screen "05-Outputs1" 480x272, template "Main_Template"
   on GenerateScreen: SetTag("DB005-HMI_Data_iScreen_Number", 5)
   TextField "TextField_ScreenName" at 76,46 size 328x30; Text 'PLC DIGITAL OUTPUTS - 1of3'
   TextField "TextField_BankLetter" at 412,50 size 64x23; Text 'BANK A'
   Button "Button_Next" at 384,227 size 92x40; TextOff 'NEXT'
      on Press: ActivateScreen("06-Outputs2", 0)
   Group "Group_DQ0.0" at 18,83 size 97x62; TextList "ON/OFF"
   Group "Group_DQ0.1" at 132,83 size 97x62; TextList "ON/OFF"
   Group "Group_DQ0.2" at 247,83 size 97x62; TextList "ON/OFF"
   Group "Group_DQ0.3" at 362,83 size 97x62; TextList "ON/OFF"
   Group "Group_DQ0.4" at 18,154 size 97x62; TextList "ON/OFF"
   Group "Group_DQ0.5" at 132,154 size 97x62; TextList "ON/OFF"
   Group "Group_DQ0.6" at 247,154 size 97x62; TextList "ON/OFF"
   Group "Group_DQ0.7" at 362,154 size 97x62; TextList "ON/OFF"
   Rectangle "Rectangle_DQ0.0" at 18,83 size 97x62
      Appearance <- "DB001-PLC_I/O_Outputs_xDQ0.0"
   TextField "Text field_DQ0.0" at 44,83 size 46x19; Text 'DQ 0.0'
   Button "Button_DQ0.0" at 30,105 size 73x32; TextOff 'Text'; TextList "ON/OFF"
      on Press: InvertBit("DB001-PLC_I/O_Outputs_xDQ0.0")
      ProcessValue <- "DB001-PLC_I/O_Outputs_xDQ0.0"
   Rectangle "Rectangle_DQ0.1" at 132,83 size 97x62
      Appearance <- "DB001-PLC_I/O_Outputs_xDQ0.1"
   TextField "Text field_DQ0.1" at 158,83 size 46x19; Text 'DQ 0.1'
   Button "Button_DQ0.1" at 144,105 size 73x32; TextOff 'Text'; TextList "ON/OFF"
      on Press: InvertBit("DB001-PLC_I/O_Outputs_xDQ0.1")
      ProcessValue <- "DB001-PLC_I/O_Outputs_xDQ0.1"
   Rectangle "Rectangle_DQ0.2" at 247,83 size 97x62
      Appearance <- "DB001-PLC_I/O_Outputs_xDQ0.2"
   TextField "Text field_DQ0.2" at 273,83 size 46x19; Text 'DQ 0.2'
   Button "Button_DQ0.2" at 259,105 size 73x32; TextOff 'Text'; TextList "ON/OFF"
      on Press: InvertBit("DB001-PLC_I/O_Outputs_xDQ0.2")
      ProcessValue <- "DB001-PLC_I/O_Outputs_xDQ0.2"
   Rectangle "Rectangle_DQ0.3" at 362,83 size 97x62
      Appearance <- "DB001-PLC_I/O_Outputs_xDQ0.3"
   TextField "Text field_DQ0.3" at 388,83 size 46x19; Text 'DQ 0.3'
   Button "Button_DQ0.3" at 374,105 size 73x32; TextOff 'Text'; TextList "ON/OFF"
      on Press: InvertBit("DB001-PLC_I/O_Outputs_xDQ0.3")
      ProcessValue <- "DB001-PLC_I/O_Outputs_xDQ0.3"
   Rectangle "Rectangle_DQ0.4" at 18,154 size 97x62
      Appearance <- "DB001-PLC_I/O_Outputs_xDQ0.4"
   TextField "Text field_DQ0.4" at 44,154 size 46x19; Text 'DQ 0.4'
   Button "Button_DQ0.4" at 30,176 size 73x32; TextOff 'Text'; TextList "ON/OFF"
      on Press: InvertBit("DB001-PLC_I/O_Outputs_xDQ0.4")
      ProcessValue <- "DB001-PLC_I/O_Outputs_xDQ0.4"
   Rectangle "Rectangle_DQ0.5" at 132,154 size 97x62
      Appearance <- "DB001-PLC_I/O_Outputs_xDQ0.5"
   TextField "Text field_DQ0.5" at 158,154 size 46x19; Text 'DQ 0.5'
   Button "Button_DQ0.5" at 144,176 size 73x32; TextOff 'Text'; TextList "ON/OFF"
      on Press: InvertBit("DB001-PLC_I/O_Outputs_xDQ0.5")
      ProcessValue <- "DB001-PLC_I/O_Outputs_xDQ0.5"
   Rectangle "Rectangle_DQ0.6" at 247,154 size 97x62
      Appearance <- "DB001-PLC_I/O_Outputs_xDQ0.6"
   TextField "Text field_DQ0.6" at 273,154 size 46x19; Text 'DQ 0.6'
   Button "Button_DQ0.6" at 259,176 size 73x32; TextOff 'Text'; TextList "ON/OFF"
      on Press: InvertBit("DB001-PLC_I/O_Outputs_xDQ0.6")
      ProcessValue <- "DB001-PLC_I/O_Outputs_xDQ0.6"
   Rectangle "Rectangle_DQ0.7" at 362,154 size 97x62
      Appearance <- "DB001-PLC_I/O_Outputs_xDQ0.7"
   TextField "Text field_DQ0.7" at 388,154 size 46x19; Text 'DQ 0.7'
   Button "Button_DQ0.7" at 374,176 size 73x32; TextOff 'Text'; TextList "ON/OFF"
      on Press: InvertBit("DB001-PLC_I/O_Outputs_xDQ0.7")
      ProcessValue <- "DB001-PLC_I/O_Outputs_xDQ0.7"

screen "08-AnalogI/O" 480x272, template "Main_Template"
   on GenerateScreen: SetTag("DB005-HMI_Data_iScreen_Number", 8)
   Button "Button_Back" at 384,227 size 92x40; TextOff 'BACK'
      on Press: function_efd93a16()
   TextField "TextField_ScreenName" at 65,46 size 351x30; Text 'PLC ANALOG INPUTS/OUTPUTS'
   Group "Group_A0" at 244,76 size 229x145; FormatPattern 9999
   Group "Group_A1" at 8,76 size 229x145; FormatPattern 9999
   TextField "Text field_A0" at 291,77 size 127x21; Text 'Analog AI-0 & AQ-0'
   TextField "Text field_A0_Input" at 279,98 size 42x17; Text 'INPUT'
   TextField "Text field_A0_Instruction" at 256,115 size 86x34; Text 'Use the connected potentiometer to change the input voltage.'
   TextField "Text field_A0_Voltage" at 280,149 size 41x14; Text 'VOLTAGE:'
   IOField "I/O field_A0_Voltage" at 281,162 size 42x21; FormatPattern 99.99; Unit  V
      ProcessValue <- "DB001-PLC_I/O_Inputs_rAI0.0_Scaled"
   TextField "Text field_A0_InRAW" at 289,181 size 24x14; Text 'RAW:'
   IOField "I/O field_A0_RAW" at 283,193 size 37x21; FormatPattern 99999
      ProcessValue <- "AI0.0"
   TextField "Text field_A0_Output" at 389,98 size 52x17; Text 'OUTPUT'
   TextField "Text field_A0_mA" at 381,127 size 19x14; Text 'mA:'
   IOField "I/O field_A0_mA" at 365,140 size 51x21; FormatPattern 99.99; Unit  mA
      ProcessValue <- "DB001-PLC_I/O_Outputs_rAQ0.0_Scaled"
   TextField "Text field_A0_OutRAW" at 379,167 size 24x14; Text 'RAW:'
   IOField "I/O field_A0_OutRAW" at 373,180 size 37x21; FormatPattern 99999
      ProcessValue <- "AQ0.0"
   TextField "Text field_A0_20" at 403,113 size 25x14; Text '20mA'
   TextField "Text field_A0_15" at 415,136 size 13x14; Text '15'
   TextField "Text field_A0_10" at 415,160 size 13x14; Text '10'
   TextField "Text field_A0_5" at 419,182 size 10x14; Text '5'
   TextField "Text field_A0_0" at 408,205 size 21x14; Text '0mA'
   Bar "Bar_A0" at 428,118 size 37x97; MinimumValue 0; MaximumValue 20
      ProcessValue <- "DB001-PLC_I/O_Outputs_rAQ0.0_Scaled"
   TextField "Text field_A1" at 55,77 size 127x21; Text 'Analog AI-1 & AQ-1'
   TextField "Text field_A1_Input" at 43,98 size 42x17; Text 'INPUT'
   TextField "Text field_A1_Instruction" at 20,115 size 86x34; Text 'Use the connected potentiometer to change the input voltage.'
   TextField "Text field_A1_Voltage" at 44,149 size 41x14; Text 'VOLTAGE:'
   IOField "I/O field_A1_Voltage" at 45,162 size 42x21; FormatPattern 99.99; Unit  V
      ProcessValue <- "DB001-PLC_I/O_Inputs_rAI0.1_Scaled"
   TextField "Text field_A1_InRAW" at 53,181 size 24x14; Text 'RAW:'
   IOField "I/O field_A1_RAW" at 47,193 size 37x21; FormatPattern 99999
      ProcessValue <- "AI0.1"
   TextField "Text field_A1_Output" at 153,98 size 52x17; Text 'OUTPUT'
   TextField "Text field_A1_mA" at 145,127 size 19x14; Text 'mA:'
   IOField "I/O field_A1_mA" at 129,140 size 51x21; FormatPattern 99.99; Unit  mA
      ProcessValue <- "DB001-PLC_I/O_Outputs_rAQ0.1_Scaled"
   TextField "Text field_A1_OutRAW" at 143,167 size 24x14; Text 'RAW:'
   IOField "I/O field_A1_OutRAW" at 137,180 size 37x21; FormatPattern 99999
      ProcessValue <- "AQ0.1"
   TextField "Text field_A1_20" at 167,113 size 25x14; Text '20mA'
   TextField "Text field_A1_15" at 179,136 size 13x14; Text '15'
   TextField "Text field_A1_10" at 179,160 size 13x14; Text '10'
   TextField "Text field_A1_5" at 183,182 size 10x14; Text '5'
   TextField "Text field_A1_0" at 172,205 size 21x14; Text '0mA'
   Bar "Bar_A1" at 192,118 size 37x97; MinimumValue 0; MaximumValue 20
      ProcessValue <- "DB001-PLC_I/O_Outputs_rAQ0.1_Scaled"

screen "03-Inputs2" 480x272, template "Main_Template"
   on GenerateScreen: SetTag("DB005-HMI_Data_iScreen_Number", 3)
   TextField "TextField_ScreenName" at 85,46 size 309x30; Text 'PLC DIGITAL INPUTS - 2of3'
   TextField "TextField_BankLetter" at 412,50 size 62x23; Text 'BANK B'
   Group "Group_DI1.0" at 73,81 size 62x63
   Group "Group_DI1.1" at 209,81 size 62x63
   Group "Group_DI1.2" at 345,81 size 62x63
   Group "Group_DI1.3" at 73,152 size 62x63
   Group "Group_DI1.4" at 209,152 size 62x64
   Group "Group_DI1.5" at 345,152 size 62x64
   TextField "Text field_DI1.0" at 83,81 size 42x19; Text 'DI 1.0'
   Circle "Circle_DI1.0" at 86,103 size 36x36
      Appearance <- "DB001-PLC_I/O_Inputs_xDI1.0"
   TextField "Text field_DI1.1" at 219,81 size 42x19; Text 'DI 1.1'
   Circle "Circle_DI1.1" at 222,103 size 36x36
      Appearance <- "DB001-PLC_I/O_Inputs_xDI1.1"
   TextField "Text field_DI1.2" at 355,81 size 42x19; Text 'DI 1.2'
   Circle "Circle_DI1.2" at 358,103 size 36x36
      Appearance <- "DB001-PLC_I/O_Inputs_xDI1.2"
   TextField "Text field_DI1.3" at 83,152 size 42x19; Text 'DI 1.3'
   Circle "Circle_DI1.3" at 86,174 size 36x36
      Appearance <- "DB001-PLC_I/O_Inputs_xDI1.3"
   TextField "Text field_DI1.4" at 219,152 size 42x19; Text 'DI 1.4'
   Circle "Circle_DI1.4" at 222,174 size 36x36
      Appearance <- "DB001-PLC_I/O_Inputs_xDI1.4"
   TextField "Text field_DI1.5" at 355,152 size 42x19; Text 'DI 1.5'
   Circle "Circle_DI1.5" at 358,174 size 36x36
      Appearance <- "DB001-PLC_I/O_Inputs_xDI1.5"
   Button "Button_Back_1" at 411,176 size 65x40; TextOff 'BACK'
      on Press: function_efd93a16()
   Button "Button_Next" at 384,227 size 92x40; TextOff 'NEXT'
      on Press: ActivateScreen("04-Inputs3", 0)

screen "06-Outputs2" 480x272, template "Main_Template"
   on GenerateScreen: SetTag("DB005-HMI_Data_iScreen_Number", 6)
   TextField "TextField_ScreenName" at 76,46 size 328x30; Text 'PLC DIGITAL OUTPUTS - 2of3'
   TextField "TextField_BankLetter" at 412,50 size 62x23; Text 'BANK B'
   Rectangle "Rectangle_DQ1.0" at 119,114 size 97x62
      Appearance <- "DB001-PLC_I/O_Outputs_xDQ1.0"
   TextField "Text field_DQ1.0" at 145,114 size 46x19; Text 'DQ 1.0'
   Button "Button_DQ1.0" at 131,136 size 73x32; TextOff 'Text'; TextList "ON/OFF"
      on Press: InvertBit("DB001-PLC_I/O_Outputs_xDQ1.0")
      ProcessValue <- "DB001-PLC_I/O_Outputs_xDQ0.0"
   Group "Group_DQ1.0" at 119,114 size 97x62; TextList "ON/OFF"
   Group "Group_DQ1.1" at 264,114 size 97x62; TextList "ON/OFF"
   Rectangle "Rectangle_DQ1.1" at 264,114 size 97x62
      Appearance <- "DB001-PLC_I/O_Outputs_xDQ1.1"
   TextField "Text field_DQ1.1" at 290,114 size 46x19; Text 'DQ 1.1'
   Button "Button_DQ1.1" at 276,136 size 73x32; TextOff 'Text'; TextList "ON/OFF"
      on Press: InvertBit("DB001-PLC_I/O_Outputs_xDQ1.1")
      ProcessValue <- "DB001-PLC_I/O_Outputs_xDQ0.1"
   Button "Button_Next" at 384,227 size 92x40; TextOff 'NEXT'
      on Press: ActivateScreen("07-Outputs3", 0)
   Button "Button_Back" at 384,181 size 92x40; TextOff 'BACK'
      on Press: function_efd93a16()

Template "Main_Template" 480x272
   GraphicView "Template_Background" at 0,0 size 480x272; Picture "HMI_Background"
   Button "Template_Button5_Blank" at 384,227 size 92x40; TextOff 'BLANK'
   Button "Template_Button1_Home" at 4,227 size 92x40; TextOff 'HOME'
      on Press: ActivateScreen("01-Home", 0)
   Button "Template_Button2_Inputs" at 99,227 size 92x40; TextOff 'INPUTS'
      on Press: ActivateScreen("02-Inputs1", 0)
   Button "Template_Button3_Outputs" at 194,227 size 92x40; TextOff 'OUTPUTS'
      on Press: ActivateScreen("05-Outputs1", 0)
   Button "Template_Button4_AnalogIO" at 289,227 size 92x40; TextOff 'ANALOG I/O'
      on Press: ActivateScreen("08-AnalogI/O", 0)
   IOField "Template_I/O field_Date" at 289,14 size 74x20; FormatPattern ????????
      ProcessValue <- "DB002-DateTime_sCustomDate_DDMMYY"
   IOField "Template_I/O field_Time" at 365,14 size 50x20; FormatPattern ?????
      ProcessValue <- "DB002-DateTime_sCustomTime_HHMM"
   GraphicView "TVET_Logo" at 8,2 size 220x44; Picture "TVET_Logo"

screen "07-Outputs3" 480x272, template "Main_Template"
   on GenerateScreen: SetTag("DB005-HMI_Data_iScreen_Number", 7)
   TextField "TextField_ScreenName" at 78,46 size 325x30; Text 'PLC IO-LINK OUTPUTS - 3of3'
   TextField "Text field_Active_Input" at 24,118 size 100x17; Text 'ACTIVE - OUTPUT'
   TextField "Text field_Active_Output" at 24,140 size 89x17; Text 'ACTIVE - INPUT'
   TextField "Text field_Port_Disabled" at 24,162 size 92x17; Text 'PORT DISABLED'
   Button "Button_Back" at 384,227 size 92x40; TextOff 'BACK'
      on Press: function_efd93a16()
   Button "Button_ConfigTL" at 338,85 size 60x56; TextOff 'CONFIG TOWER LIGHT'
      on Press: ActivateScreen("09-TowerLight_Config", 0)
   TextField "Text field_X01" at 168,81 size 28x19; Text 'X01'
   Group "Group_X01" at 152,81 size 62x63
   Group "Group_X02" at 268,81 size 62x63
   Group "Group_X03" at 152,152 size 62x63
   Group "Group_X04" at 268,152 size 62x63
   TextField "Text field_X02" at 284,81 size 28x19; Text 'X02'
   TextField "Text field_X03" at 168,152 size 28x19; Text 'X03'
   TextField "Text field_X04" at 284,152 size 28x19; Text 'X04'

screen "04-Inputs3" 480x272, template "Main_Template"
   on GenerateScreen: SetTag("DB005-HMI_Data_iScreen_Number", 4)
   Button "Button_Back" at 384,227 size 92x40; TextOff 'BACK'
      on Press: function_efd93a16()
   TextField "TextField_ScreenName" at 87,46 size 306x30; Text 'PLC IO-LINK INPUTS - 3of3'
   TextField "Text field_Active_Input" at 24,118 size 89x17; Text 'ACTIVE - INPUT'
   TextField "Text field_Active_Output" at 24,140 size 100x17; Text 'ACTIVE - OUTPUT'
   TextField "Text field_Port_Disabled" at 24,162 size 92x17; Text 'PORT DISABLED'
   TextField "Text field_X02" at 284,81 size 28x19; Text 'X02'
   TextField "Text field_X03" at 168,152 size 28x19; Text 'X03'
   TextField "Text field_X04" at 284,152 size 28x19; Text 'X04'
   TextField "Text field_X01" at 168,81 size 28x19; Text 'X01'
   Group "Group_X01" at 152,81 size 62x63
   Group "Group_X02" at 268,81 size 62x63
   Group "Group_X03" at 152,152 size 62x63
   Group "Group_X04" at 268,152 size 62x63

screen "09-TowerLight_Config" 480x272, template "Main_Template"
   on GenerateScreen: SetTag("DB005-HMI_Data_iScreen_Number", 9)
   Button "Button_Back" at 384,227 size 92x40; TextOff 'BACK'
      on Press: function_efd93a16()
   TextField "TextField_ScreenName" at 60,46 size 360x30; Text 'IO-LINK_TOWERLIGHT_CONFIG'
   Button "Button_Save_Config" at 376,160 size 53x43; TextOff 'SAVE CONFIG'
      on Press: InvertBit("DB005-HMI_Data_TowerLight_xSave_Config")
      Appearance <- "DB005-HMI_Data_TowerLight_xSave_Config"
      on Release: InvertBit("DB005-HMI_Data_TowerLight_xSave_Config")
   TextField "Text field_Segment1" at 45,81 size 58x17; Text 'SEGMENT1'
   TextField "Text field_Seg1_Animate" at 24,102 size 40x14; Text 'ANIMATE:'
   SymbolicIOField "Symbolic I/O field_Seg1_Animate" at 66,101 size 64x16; TextOff '0'; TextOn '1'; TextList "Animate"
      ProcessValue <- "DB005-HMI_Data_TowerLight_Segment1_iAnimate"
   TextField "Text field_Seg1_Colour1" at 24,126 size 42x14; Text 'COLOUR1:'
   SymbolicIOField "Symbolic I/O field_Seg1_Colour1" at 66,125 size 64x16; TextOff '0'; TextOn '1'; TextList "Colour1"
      ProcessValue <- "DB005-HMI_Data_TowerLight_Segment1_iColour1"
   TextField "Text field_Seg1_Colour2" at 24,150 size 42x14; Text 'COLOUR2:'
   SymbolicIOField "Symbolic I/O field_Seg1_Colour2" at 66,149 size 64x16; TextOff '0'; TextOn '1'; TextList "Colour2"
      ProcessValue <- "DB005-HMI_Data_TowerLight_Segment1_iColour2"
   TextField "Text field_Seg1_Speed" at 24,174 size 28x14; Text 'SPEED:'
   SymbolicIOField "Symbolic I/O field_Seg1_Speed" at 66,173 size 64x16; TextOff '0'; TextOn '1'; TextList "Speed"
      ProcessValue <- "DB005-HMI_Data_TowerLight_Segment1_iSpeed"
   TextField "Text field_Seg1_Colour_Width_Percent" at 24,198 size 39x14; Text 'CLR W%:'
   TextField "Text field_Seg1_1-100" at 24,205 size 29x14; Text '(1-100)'
   IOField "I/O field_Seg1_Colour_Width_Percent" at 66,197 size 64x16; FormatPattern 999
      ProcessValue <- "DB005-HMI_Data_TowerLight_Segment1_iClrWidth%"
   TextField "Text field_Segment2" at 153,81 size 58x17; Text 'SEGMENT2'
   TextField "Text field_Seg2_Animate" at 132,102 size 40x14; Text 'ANIMATE:'
   SymbolicIOField "Symbolic I/O field_Seg2_Animate" at 174,101 size 64x16; TextOff '0'; TextOn '1'; TextList "Animate"
      ProcessValue <- "DB005-HMI_Data_TowerLight_Segment2_iAnimate"
   TextField "Text field_Seg2_Colour1" at 132,126 size 42x14; Text 'COLOUR1:'
   SymbolicIOField "Symbolic I/O field_Seg2_Colour1" at 174,125 size 64x16; TextOff '0'; TextOn '1'; TextList "Colour1"
      ProcessValue <- "DB005-HMI_Data_TowerLight_Segment2_iColour1"
   TextField "Text field_Seg2_Colour2" at 132,150 size 42x14; Text 'COLOUR2:'
   SymbolicIOField "Symbolic I/O field_Seg2_Colour2" at 174,149 size 64x16; TextOff '0'; TextOn '1'; TextList "Colour2"
      ProcessValue <- "DB005-HMI_Data_TowerLight_Segment2_iColour2"
   TextField "Text field_Seg2_Speed" at 132,174 size 28x14; Text 'SPEED:'
   SymbolicIOField "Symbolic I/O field_Seg2_Speed" at 174,173 size 64x16; TextOff '0'; TextOn '1'; TextList "Speed"
      ProcessValue <- "DB005-HMI_Data_TowerLight_Segment2_iSpeed"
   TextField "Text field_Seg2_Colour_Width_Percent" at 132,198 size 39x14; Text 'CLR W%:'
   TextField "Text field_Seg2_1-100" at 132,205 size 29x14; Text '(1-100)'
   IOField "I/O field_Seg2_Colour_Width_Percent" at 174,197 size 64x16; FormatPattern 999
      ProcessValue <- "DB005-HMI_Data_TowerLight_Segment2_iClrWidth%"
   TextField "Text field_Segment3" at 261,81 size 58x17; Text 'SEGMENT3'
   TextField "Text field_Seg3_Animate" at 240,102 size 40x14; Text 'ANIMATE:'
   SymbolicIOField "Symbolic I/O field_Seg3_Animate" at 282,101 size 64x16; TextOff '0'; TextOn '1'; TextList "Animate"
      ProcessValue <- "DB005-HMI_Data_TowerLight_Segment3_iAnimate"
   TextField "Text field_Seg3_Colour1" at 240,126 size 42x14; Text 'COLOUR1:'
   SymbolicIOField "Symbolic I/O field_Seg3_Colour1" at 282,125 size 64x16; TextOff '0'; TextOn '1'; TextList "Colour1"
      ProcessValue <- "DB005-HMI_Data_TowerLight_Segment3_iColour1"
   TextField "Text field_Seg3_Colour2" at 240,150 size 42x14; Text 'COLOUR2:'
   SymbolicIOField "Symbolic I/O field_Seg3_Colour2" at 282,149 size 64x16; TextOff '0'; TextOn '1'; TextList "Colour2"
      ProcessValue <- "DB005-HMI_Data_TowerLight_Segment3_iColour2"
   TextField "Text field_Seg3_Speed" at 240,174 size 28x14; Text 'SPEED:'
   SymbolicIOField "Symbolic I/O field_Seg3_Speed" at 282,173 size 64x16; TextOff '0'; TextOn '1'; TextList "Speed"
      ProcessValue <- "DB005-HMI_Data_TowerLight_Segment3_iSpeed"
   TextField "Text field_Seg3_Colour_Width_Percent" at 240,198 size 39x14; Text 'CLR W%:'
   TextField "Text field_Seg3_1-100" at 240,205 size 29x14; Text '(1-100)'
   IOField "I/O field_Seg3_Colour_Width_Percent" at 282,197 size 64x16; FormatPattern 999
      ProcessValue <- "DB005-HMI_Data_TowerLight_Segment3_iClrWidth%"
   TextField "Text field_Audible" at 377,81 size 48x17; Text 'AUDIBLE'
   TextField "Text field_Volume" at 348,102 size 37x14; Text 'VOLUME:'
   SymbolicIOField "Symbolic I/O field_Volume" at 390,101 size 64x16; TextOff '0'; TextOn '1'; TextList "Volume"
      ProcessValue <- "DB005-HMI_Data_TowerLight_Audible_iVolume"
   TextField "Text field_Type" at 348,126 size 25x14; Text 'TYPE:'
   SymbolicIOField "Symbolic I/O field_Type" at 390,125 size 64x16; TextOff '0'; TextOn '1'; TextList "Type"
      ProcessValue <- "DB005-HMI_Data_TowerLight_Audible_iType"
*)